(* Logix 5000 project; controller Almacen_1 vendor 1 type 14 code 235 rev 36.11; software revision 36.00; part 2 of 2 *)
(* tags used below, declared in another part *)
   Contador_Salida_Conveyor : COUNTER;
   End_Conveyor_Rutine : BOOL;
   Start_Conveyor_1 : BOOL;
   Start_Rutine : BOOL;
   Stop_Conveyor_1 : BOOL;
   tag_switch : BOOL;
   tag_switch2 : BOOL;
   tag_switch3 : BOOL;
   Tag_switch4 : BOOL;
   tag_switch5 : BOOL;
   tag_switch6 : BOOL;
   tag_timer_piston : BOOL;
   tag_timer_piston2 : BOOL;
   Timer1_Cambio_Direccion_CNC : TIMER;
   Timer2 : TIMER;
   Timer3_Piston_Marcadora_OFF : TIMER;
   Timer4_Piston_Camara_ON : TIMER;
   Timer5_Piston_Camara_OFF : TIMER;
   Timer6_Cambio_Direccion_Almacen : TIMER;
   Timer7_Sensor_Entrada_Salida : TIMER;
   Timer8_Stop_Conveyor : TIMER;
   Timer9_Piston_Salida : TIMER;
   At_Pos_Alm_1 : DINT;
   In_Pos_Alm_1 : DINT;
   PosicionAlmacen : DINT;
   Start_Kinetix_Alm_1 : DINT;
   Start_Motor_Alm_1 : BOOL;
   To_Pos_Alm_1 : DINT;
(* MainProgram, continued *)

ROUTINE Camara_t   (* ladder *)
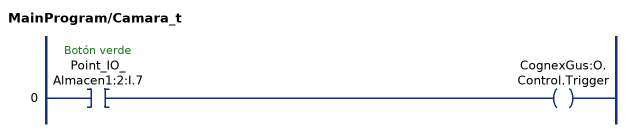
   0: XIC(Point_IO_Almacen1:2:I.7)OTE(CognexGus:O.Control.Trigger);
END_ROUTINE

ROUTINE MainRoutine   (* ladder *)
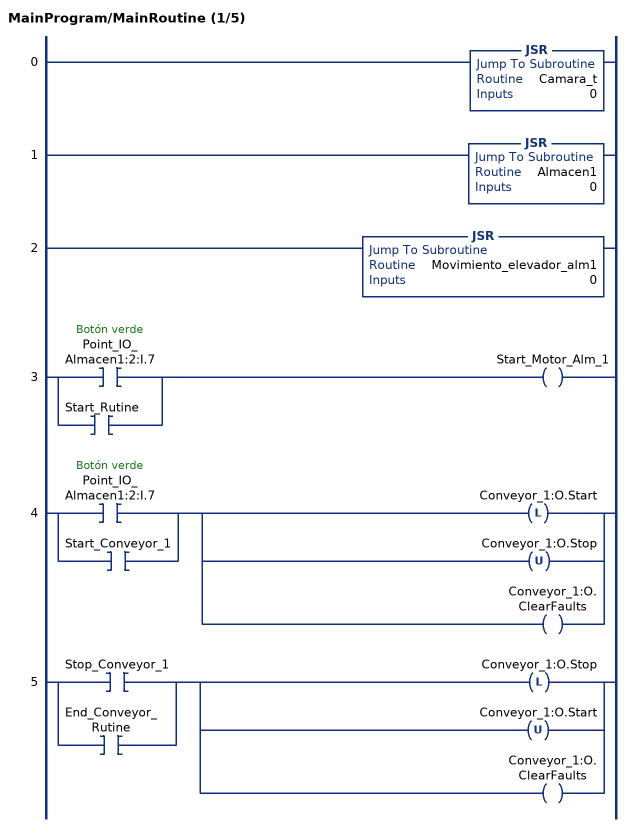
   0: JSR(Camara_t,0);
   1: JSR(Almacen1,0);
   2: JSR(Movimiento_elevador_alm1,0);
   3: [XIC(Point_IO_Almacen1:2:I.7) ,XIC(Start_Rutine) ]OTE(Start_Motor_Alm_1);
   4: [XIC(Point_IO_Almacen1:2:I.7) ,XIC(Start_Conveyor_1) ][OTL(Conveyor_1:O.Start) ,OTU(Conveyor_1:O.Stop) ,OTE(Conveyor_1:O.ClearFaults) ];
   5: [XIC(Stop_Conveyor_1) ,XIC(End_Conveyor_Rutine) ][OTL(Conveyor_1:O.Stop) ,OTU(Conveyor_1:O.Start) ,OTE(Conveyor_1:O.ClearFaults) ];
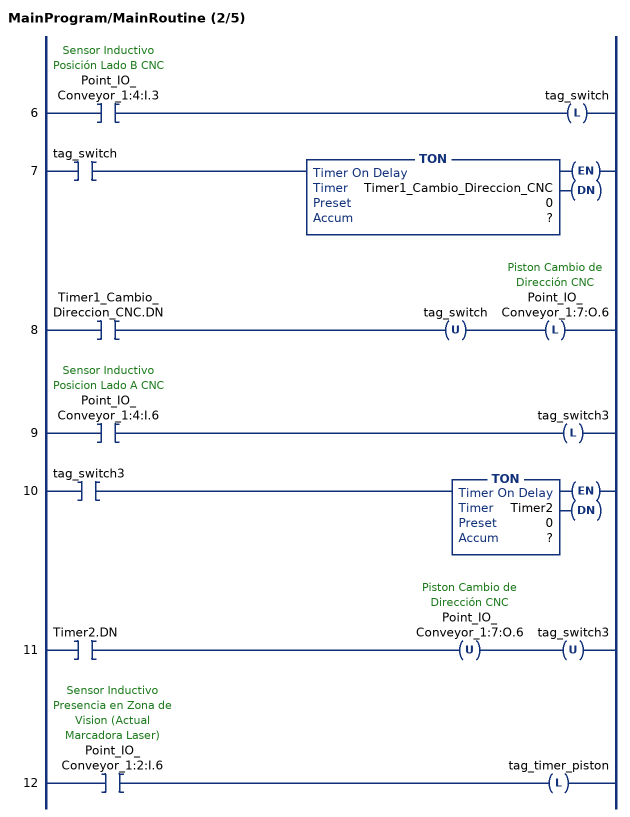
   6: XIC(Point_IO_Conveyor_1:4:I.3)OTL(tag_switch);
   7: XIC(tag_switch)TON(Timer1_Cambio_Direccion_CNC,?,?);
   8: XIC(Timer1_Cambio_Direccion_CNC.DN)OTU(tag_switch)OTL(Point_IO_Conveyor_1:7:O.6);
   9: XIC(Point_IO_Conveyor_1:4:I.6)OTL(tag_switch3);
   10: XIC(tag_switch3)TON(Timer2,?,?);
   11: XIC(Timer2.DN)OTU(Point_IO_Conveyor_1:7:O.6)OTU(tag_switch3);
   12: XIC(Point_IO_Conveyor_1:2:I.6)OTL(tag_timer_piston);
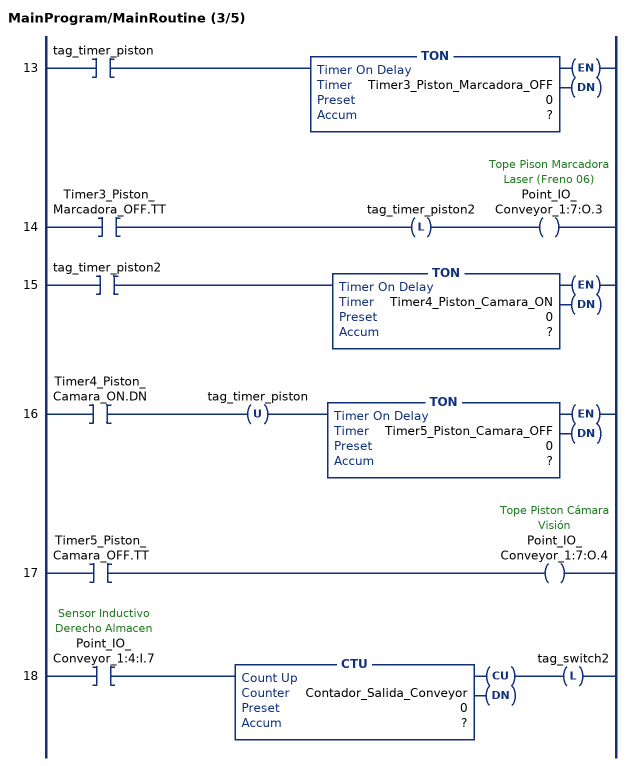
   13: XIC(tag_timer_piston)TON(Timer3_Piston_Marcadora_OFF,?,?);
   14: XIC(Timer3_Piston_Marcadora_OFF.TT)OTL(tag_timer_piston2)OTE(Point_IO_Conveyor_1:7:O.3);
   15: XIC(tag_timer_piston2)TON(Timer4_Piston_Camara_ON,?,?);
   16: XIC(Timer4_Piston_Camara_ON.DN)OTU(tag_timer_piston)TON(Timer5_Piston_Camara_OFF,?,?);
   17: XIC(Timer5_Piston_Camara_OFF.TT)OTE(Point_IO_Conveyor_1:7:O.4);
   18: XIC(Point_IO_Conveyor_1:4:I.7)CTU(Contador_Salida_Conveyor,?,?)OTL(tag_switch2);
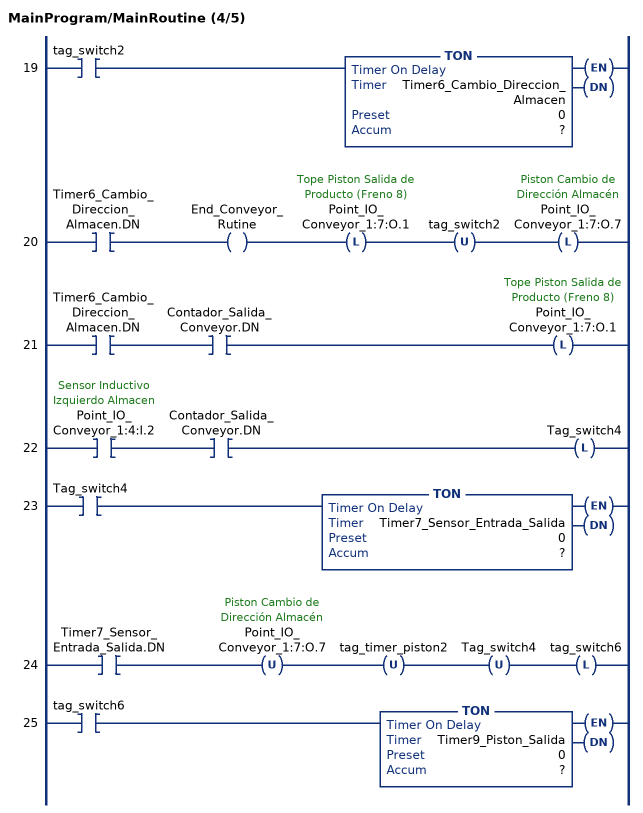
   19: XIC(tag_switch2)TON(Timer6_Cambio_Direccion_Almacen,?,?);
   20: XIC(Timer6_Cambio_Direccion_Almacen.DN)OTE(End_Conveyor_Rutine)OTL(Point_IO_Conveyor_1:7:O.1)OTU(tag_switch2)OTL(Point_IO_Conveyor_1:7:O.7);
   21: XIC(Timer6_Cambio_Direccion_Almacen.DN)XIC(Contador_Salida_Conveyor.DN)OTL(Point_IO_Conveyor_1:7:O.1);
   22: XIC(Point_IO_Conveyor_1:4:I.2)XIC(Contador_Salida_Conveyor.DN)OTL(Tag_switch4);
   23: XIC(Tag_switch4)TON(Timer7_Sensor_Entrada_Salida,?,?);
   24: XIC(Timer7_Sensor_Entrada_Salida.DN)OTU(Point_IO_Conveyor_1:7:O.7)OTU(tag_timer_piston2)OTU(Tag_switch4)OTL(tag_switch6);
   25: XIC(tag_switch6)TON(Timer9_Piston_Salida,?,?);
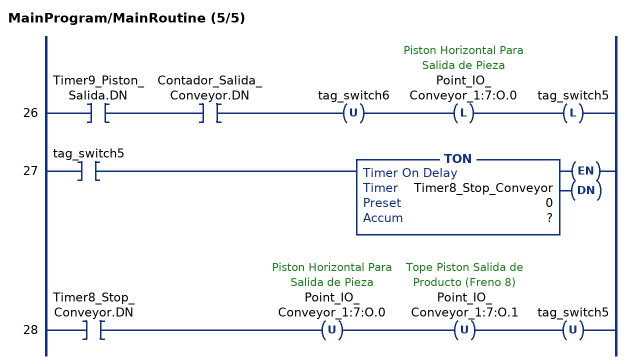
   26: XIC(Timer9_Piston_Salida.DN)XIC(Contador_Salida_Conveyor.DN)OTU(tag_switch6)OTL(Point_IO_Conveyor_1:7:O.0)OTL(tag_switch5);
   27: XIC(tag_switch5)TON(Timer8_Stop_Conveyor,?,?);
   28: XIC(Timer8_Stop_Conveyor.DN)OTU(Point_IO_Conveyor_1:7:O.0)OTU(Point_IO_Conveyor_1:7:O.1)OTU(tag_switch5);
END_ROUTINE

ROUTINE Movimiento_elevador_alm1   (* ladder *)
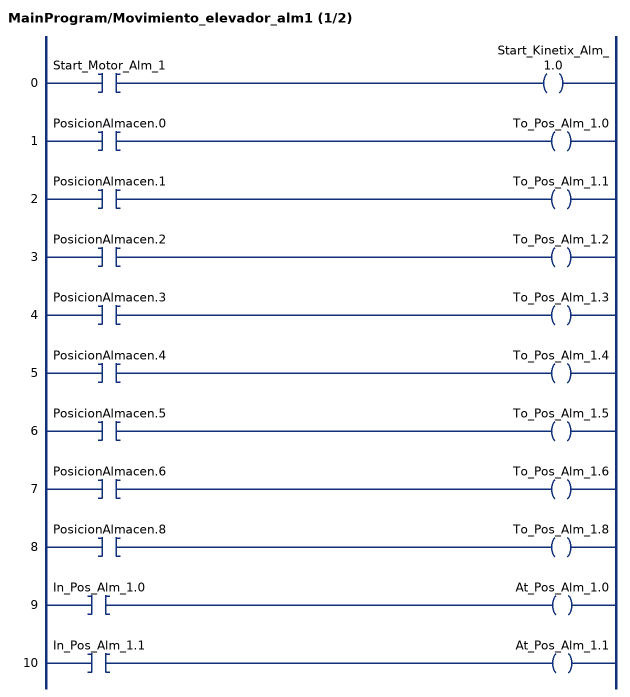
   0: XIC(Start_Motor_Alm_1)OTE(Start_Kinetix_Alm_1.0);
   1: XIC(PosicionAlmacen.0)OTE(To_Pos_Alm_1.0);
   2: XIC(PosicionAlmacen.1)OTE(To_Pos_Alm_1.1);
   3: XIC(PosicionAlmacen.2)OTE(To_Pos_Alm_1.2);
   4: XIC(PosicionAlmacen.3)OTE(To_Pos_Alm_1.3);
   5: XIC(PosicionAlmacen.4)OTE(To_Pos_Alm_1.4);
   6: XIC(PosicionAlmacen.5)OTE(To_Pos_Alm_1.5);
   7: XIC(PosicionAlmacen.6)OTE(To_Pos_Alm_1.6);
   8: XIC(PosicionAlmacen.8)OTE(To_Pos_Alm_1.8);
   9: XIC(In_Pos_Alm_1.0)OTE(At_Pos_Alm_1.0);
   10: XIC(In_Pos_Alm_1.1)OTE(At_Pos_Alm_1.1);
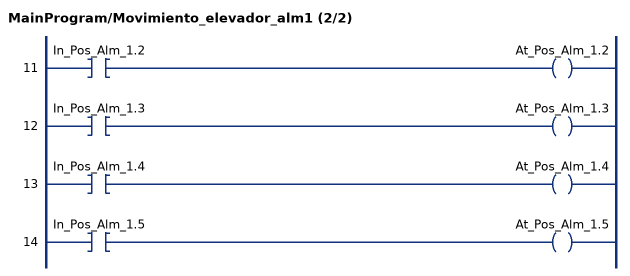
   11: XIC(In_Pos_Alm_1.2)OTE(At_Pos_Alm_1.2);
   12: XIC(In_Pos_Alm_1.3)OTE(At_Pos_Alm_1.3);
   13: XIC(In_Pos_Alm_1.4)OTE(At_Pos_Alm_1.4);
   14: XIC(In_Pos_Alm_1.5)OTE(At_Pos_Alm_1.5);
END_ROUTINE
END_PROGRAM

PROGRAM SafetyProgram   (* main routine MainRoutine, safety *)

ROUTINE MainRoutine   (* ladder *)
END_ROUTINE
END_PROGRAM
